   t[8557] := 3_855_850_566;
   t[8558] := 855_950_567;
   t[8559] := 1_856_050_568;
   t[8560] := 2_856_150_569;
   t[8561] := 2_856_250_570;
   t[8562] := 2_856_350_571;
   t[8563] := 1_856_450_572;
   t[8564] := 1_856_550_573;
   t[8565] := 2_856_650_574;
   t[8566] := 2_856_750_575;
   t[8567] := 3_856_850_576;
   t[8568] := 856_950_577;
   t[8569] := 1_857_050_578;
   t[8570] := 1_857_150_579;
   t[8571] := 1_857_250_580;
   t[8572] := 1_857_350_581;
   t[8573] := 2_857_450_582;
   t[8574] := 2_857_550_583;
   t[8575] := 2_857_650_584;
   t[8576] := 3_857_750_585;
   t[8577] := 3_857_850_586;
   t[8578] := 1_857_950_587;
   t[8579] := 1_858_050_588;
   t[8580] := 3_858_150_589;
   t[8581] := 1_858_250_590;
   t[8582] := 3_858_350_591;
   t[8583] := 1_858_450_592;
   t[8584] := 3_858_550_593;
   t[8585] := 858_650_594;
   t[8586] := 858_750_595;
   t[8587] := 1_858_850_596;
   t[8588] := 1_858_950_597;
   t[8589] := 2_859_050_598;
   t[8590] := 1_859_150_599;
   t[8591] := 3_859_250_600;
   t[8592] := 2_859_350_601;
   t[8593] := 859_450_602;
   t[8594] := 859_550_603;
   t[8595] := 1_859_650_604;
   t[8596] := 3_859_750_605;
   t[8597] := 859_850_606;
   t[8598] := 859_950_607;
   t[8599] := 2_860_050_608;
   t[8600] := 3_860_150_609;
   t[8601] := 1_860_250_610;
   t[8602] := 1_860_350_611;
   t[8603] := 2_860_450_612;
   t[8604] := 2_860_550_613;
   t[8605] := 3_860_650_614;
   t[8606] := 3_860_750_615;
   t[8607] := 3_860_850_616;
   t[8608] := 860_950_617;
   t[8609] := 3_861_050_618;
   t[8610] := 861_150_619;
   t[8611] := 861_250_620;
   t[8612] := 2_861_350_621;
   t[8613] := 2_861_450_622;
   t[8614] := 3_861_550_623;
   t[8615] := 2_861_650_624;
   t[8616] := 861_750_625;
   t[8617] := 3_861_850_626;
   t[8618] := 861_950_627;
   t[8619] := 1_862_050_628;
   t[8620] := 1_862_150_629;
   t[8621] := 3_862_250_630;
   t[8622] := 2_862_350_631;
   t[8623] := 3_862_450_632;
   t[8624] := 2_862_550_633;
   t[8625] := 3_862_650_634;
   t[8626] := 3_862_750_635;
   t[8627] := 862_850_636;
   t[8628] := 2_862_950_637;
   t[8629] := 2_863_050_638;
   t[8630] := 863_150_639;
   t[8631] := 3_863_250_640;
   t[8632] := 1_863_350_641;
   t[8633] := 3_863_450_642;
   t[8634] := 3_863_550_643;
   t[8635] := 1_863_650_644;
   t[8636] := 3_863_750_645;
   t[8637] := 1_863_850_646;
   t[8638] := 863_950_647;
   t[8639] := 2_864_050_648;
   t[8640] := 1_864_150_649;
   t[8641] := 2_864_250_650;
   t[8642] := 864_350_651;
   t[8643] := 864_450_652;
   t[8644] := 2_864_550_653;
   t[8645] := 1_864_650_654;
   t[8646] := 3_864_750_655;
   t[8647] := 3_864_850_656;
   t[8648] := 2_864_950_657;
   t[8649] := 865_050_658;
   t[8650] := 1_865_150_659;
   t[8651] := 3_865_250_660;
   t[8652] := 2_865_350_661;
   t[8653] := 865_450_662;
   t[8654] := 3_865_550_663;
   t[8655] := 865_650_664;
   t[8656] := 865_750_665;
   t[8657] := 1_865_850_666;
   t[8658] := 2_865_950_667;
   t[8659] := 3_866_050_668;
   t[8660] := 866_150_669;
   t[8661] := 1_866_250_670;
   t[8662] := 3_866_350_671;
   t[8663] := 2_866_450_672;
   t[8664] := 866_550_673;
   t[8665] := 3_866_650_674;
   t[8666] := 1_866_750_675;
   t[8667] := 1_866_850_676;
   t[8668] := 2_866_950_677;
   t[8669] := 2_867_050_678;
   t[8670] := 3_867_150_679;
   t[8671] := 2_867_250_680;
   t[8672] := 867_350_681;
   t[8673] := 867_450_682;
   t[8674] := 1_867_550_683;
   t[8675] := 867_650_684;
   t[8676] := 2_867_750_685;
   t[8677] := 2_867_850_686;
   t[8678] := 3_867_950_687;
   t[8679] := 3_868_050_688;
   t[8680] := 868_150_689;
   t[8681] := 1_868_250_690;
   t[8682] := 1_868_350_691;
   t[8683] := 2_868_450_692;
   t[8684] := 3_868_550_693;
   t[8685] := 868_650_694;
   t[8686] := 868_750_695;
   t[8687] := 1_868_850_696;
   t[8688] := 2_868_950_697;
   t[8689] := 2_869_050_698;
   t[8690] := 869_150_699;
   t[8691] := 3_869_250_700;
   t[8692] := 1_869_350_701;
   t[8693] := 869_450_702;
   t[8694] := 1_869_550_703;
   t[8695] := 1_869_650_704;
   t[8696] := 2_869_750_705;
   t[8697] := 2_869_850_706;
   t[8698] := 3_869_950_707;
   t[8699] := 3_870_050_708;
   t[8700] := 870_150_709;
   t[8701] := 870_250_710;
   t[8702] := 1_870_350_711;
   t[8703] := 3_870_450_712;
   t[8704] := 3_870_550_713;
   t[8705] := 1_870_650_714;
   t[8706] := 870_750_715;
   t[8707] := 2_870_850_716;
   t[8708] := 2_870_950_717;
   t[8709] := 2_871_050_718;
   t[8710] := 3_871_150_719;
   t[8711] := 3_871_250_720;
   t[8712] := 1_871_350_721;
   t[8713] := 1_871_450_722;
   t[8714] := 2_871_550_723;
   t[8715] := 2_871_650_724;
   t[8716] := 2_871_750_725;
   t[8717] := 1_871_850_726;
   t[8718] := 3_871_950_727;
   t[8719] := 2_872_050_728;
   t[8720] := 872_150_729;
   t[8721] := 872_250_730;
   t[8722] := 1_872_350_731;
   t[8723] := 2_872_450_732;
   t[8724] := 2_872_550_733;
   t[8725] := 872_650_734;
   t[8726] := 3_872_750_735;
   t[8727] := 1_872_850_736;
   t[8728] := 872_950_737;
   t[8729] := 2_873_050_738;
   t[8730] := 2_873_150_739;
   t[8731] := 873_250_740;
   t[8732] := 873_350_741;
   t[8733] := 1_873_450_742;
   t[8734] := 3_873_550_743;
   t[8735] := 873_650_744;
   t[8736] := 2_873_750_745;
   t[8737] := 1_873_850_746;
   t[8738] := 3_873_950_747;
   t[8739] := 2_874_050_748;
   t[8740] := 874_150_749;
   t[8741] := 1_874_250_750;
   t[8742] := 1_874_350_751;
   t[8743] := 3_874_450_752;
   t[8744] := 2_874_550_753;
   t[8745] := 874_650_754;
   t[8746] := 874_750_755;
   t[8747] := 1_874_850_756;
   t[8748] := 2_874_950_757;
   t[8749] := 3_875_050_758;
   t[8750] := 875_150_759;
   t[8751] := 875_250_760;
   t[8752] := 2_875_350_761;
   t[8753] := 2_875_450_762;
   t[8754] := 3_875_550_763;
   t[8755] := 2_875_650_764;
   t[8756] := 875_750_765;
   t[8757] := 1_875_850_766;
   t[8758] := 1_875_950_767;
   t[8759] := 3_876_050_768;
   t[8760] := 876_150_769;
   t[8761] := 1_876_250_770;
   t[8762] := 876_350_771;
   t[8763] := 2_876_450_772;
   t[8764] := 2_876_550_773;
   t[8765] := 876_650_774;
   t[8766] := 3_876_750_775;
   t[8767] := 876_850_776;
   t[8768] := 3_876_950_777;
   t[8769] := 1_877_050_778;
   t[8770] := 1_877_150_779;
   t[8771] := 2_877_250_780;
   t[8772] := 3_877_350_781;
   t[8773] := 877_450_782;
   t[8774] := 2_877_550_783;
   t[8775] := 2_877_650_784;
   t[8776] := 877_750_785;
   t[8777] := 2_877_850_786;
   t[8778] := 877_950_787;
   t[8779] := 3_878_050_788;
   t[8780] := 1_878_150_789;
   t[8781] := 2_878_250_790;
   t[8782] := 2_878_350_791;
   t[8783] := 878_450_792;
   t[8784] := 3_878_550_793;
   t[8785] := 878_650_794;
   t[8786] := 3_878_750_795;
   t[8787] := 1_878_850_796;
   t[8788] := 1_878_950_797;
   t[8789] := 2_879_050_798;
   t[8790] := 3_879_150_799;
   t[8791] := 879_250_800;
   t[8792] := 879_350_801;
   t[8793] := 879_450_802;
   t[8794] := 879_550_803;
   t[8795] := 879_650_804;
   t[8796] := 879_750_805;
   t[8797] := 879_850_806;
   t[8798] := 879_950_807;
   t[8799] := 880_050_808;
   t[8800] := 880_150_809;
   t[8801] := 880_250_810;
   t[8802] := 1_880_350_811;
   t[8803] := 2_880_450_812;
   t[8804] := 3_880_550_813;
   t[8805] := 880_650_814;
   t[8806] := 880_750_815;
   t[8807] := 880_850_816;
   t[8808] := 1_880_950_817;
   t[8809] := 1_881_050_818;
   t[8810] := 3_881_150_819;
   t[8811] := 3_881_250_820;
   t[8812] := 1_881_350_821;
   t[8813] := 2_881_450_822;
   t[8814] := 3_881_550_823;
   t[8815] := 881_650_824;
   t[8816] := 881_750_825;
   t[8817] := 881_850_826;
   t[8818] := 3_881_950_827;
   t[8819] := 3_882_050_828;
   t[8820] := 882_150_829;
   t[8821] := 882_250_830;
   t[8822] := 1_882_350_831;
   t[8823] := 882_450_832;
   t[8824] := 1_882_550_833;
   t[8825] := 1_882_650_834;
   t[8826] := 2_882_750_835;
   t[8827] := 1_882_850_836;
   t[8828] := 3_882_950_837;
   t[8829] := 3_883_050_838;
   t[8830] := 883_150_839;
   t[8831] := 883_250_840;
   t[8832] := 1_883_350_841;
   t[8833] := 2_883_450_842;
   t[8834] := 3_883_550_843;
   t[8835] := 883_650_844;
   t[8836] := 883_750_845;
   t[8837] := 2_883_850_846;
   t[8838] := 2_883_950_847;
   t[8839] := 3_884_050_848;
   t[8840] := 3_884_150_849;
   t[8841] := 1_884_250_850;
   t[8842] := 1_884_350_851;
   t[8843] := 2_884_450_852;
   t[8844] := 1_884_550_853;
   t[8845] := 3_884_650_854;
   t[8846] := 2_884_750_855;
   t[8847] := 884_850_856;
   t[8848] := 884_950_857;
   t[8849] := 2_885_050_858;
   t[8850] := 3_885_150_859;
   t[8851] := 1_885_250_860;
   t[8852] := 1_885_350_861;
   t[8853] := 3_885_450_862;
   t[8854] := 3_885_550_863;
   t[8855] := 885_650_864;
   t[8856] := 1_885_750_865;
   t[8857] := 2_885_850_866;
   t[8858] := 3_885_950_867;
   t[8859] := 886_050_868;
   t[8860] := 886_150_869;
   t[8861] := 886_250_870;
   t[8862] := 886_350_871;
   t[8863] := 1_886_450_872;
   t[8864] := 1_886_550_873;
   t[8865] := 1_886_650_874;
   t[8866] := 1_886_750_875;
   t[8867] := 1_886_850_876;
   t[8868] := 1_886_950_877;
   t[8869] := 887_050_878;
   t[8870] := 887_150_879;
   t[8871] := 2_887_250_880;
   t[8872] := 2_887_350_881;
   t[8873] := 887_450_882;
   t[8874] := 887_550_883;
   t[8875] := 2_887_650_884;
   t[8876] := 1_887_750_885;
   t[8877] := 1_887_850_886;
   t[8878] := 887_950_887;
   t[8879] := 2_888_050_888;
   t[8880] := 2_888_150_889;
   t[8881] := 888_250_890;
   t[8882] := 888_350_891;
   t[8883] := 2_888_450_892;
   t[8884] := 3_888_550_893;
   t[8885] := 3_888_650_894;
   t[8886] := 888_750_895;
   t[8887] := 3_888_850_896;
   t[8888] := 1_888_950_897;
   t[8889] := 1_889_050_898;
   t[8890] := 3_889_150_899;
   t[8891] := 889_250_900;
   t[8892] := 889_350_901;
   t[8893] := 1_889_450_902;
   t[8894] := 2_889_550_903;
   t[8895] := 889_650_904;
   t[8896] := 889_750_905;
   t[8897] := 2_889_850_906;
   t[8898] := 2_889_950_907;
   t[8899] := 890_050_908;
   t[8900] := 3_890_150_909;
   t[8901] := 1_890_250_910;
   t[8902] := 1_890_350_911;
   t[8903] := 2_890_450_912;
   t[8904] := 2_890_550_913;
   t[8905] := 890_650_914;
   t[8906] := 890_750_915;
   t[8907] := 1_890_850_916;
   t[8908] := 1_890_950_917;
   t[8909] := 3_891_050_918;
   t[8910] := 1_891_150_919;
   t[8911] := 3_891_250_920;
   t[8912] := 1_891_350_921;
   t[8913] := 1_891_450_922;
   t[8914] := 3_891_550_923;
   t[8915] := 3_891_650_924;
   t[8916] := 891_750_925;
   t[8917] := 2_891_850_926;
   t[8918] := 1_891_950_927;
   t[8919] := 3_892_050_928;
   t[8920] := 2_892_150_929;
   t[8921] := 3_892_250_930;
   t[8922] := 1_892_350_931;
   t[8923] := 892_450_932;
   t[8924] := 2_892_550_933;
   t[8925] := 2_892_650_934;
   t[8926] := 892_750_935;
   t[8927] := 1_892_850_936;
   t[8928] := 2_892_950_937;
   t[8929] := 893_050_938;
   t[8930] := 893_150_939;
   t[8931] := 2_893_250_940;
   t[8932] := 2_893_350_941;
   t[8933] := 893_450_942;
   t[8934] := 3_893_550_943;
   t[8935] := 1_893_650_944;
   t[8936] := 1_893_750_945;
   t[8937] := 2_893_850_946;
   t[8938] := 2_893_950_947;
   t[8939] := 3_894_050_948;
   t[8940] := 894_150_949;
   t[8941] := 1_894_250_950;
   t[8942] := 2_894_350_951;
   t[8943] := 3_894_450_952;
   t[8944] := 894_550_953;
   t[8945] := 894_650_954;
   t[8946] := 894_750_955;
   t[8947] := 894_850_956;
   t[8948] := 1_894_950_957;
   t[8949] := 1_895_050_958;
   t[8950] := 2_895_150_959;
   t[8951] := 3_895_250_960;
   t[8952] := 895_350_961;
   t[8953] := 895_450_962;
   t[8954] := 3_895_550_963;
   t[8955] := 1_895_650_964;
   t[8956] := 1_895_750_965;
   t[8957] := 3_895_850_966;
   t[8958] := 3_895_950_967;
   t[8959] := 1_896_050_968;
   t[8960] := 1_896_150_969;
   t[8961] := 2_896_250_970;
   t[8962] := 2_896_350_971;
   t[8963] := 3_896_450_972;
   t[8964] := 896_550_973;
   t[8965] := 2_896_650_974;
   t[8966] := 3_896_750_975;
   t[8967] := 1_896_850_976;
   t[8968] := 1_896_950_977;
   t[8969] := 2_897_050_978;
   t[8970] := 3_897_150_979;
   t[8971] := 3_897_250_980;
   t[8972] := 897_350_981;
   t[8973] := 1_897_450_982;
   t[8974] := 2_897_550_983;
   t[8975] := 1_897_650_984;
   t[8976] := 1_897_750_985;
   t[8977] := 1_897_850_986;
   t[8978] := 1_897_950_987;
   t[8979] := 898_050_988;
   t[8980] := 1_898_150_989;
   t[8981] := 1_898_250_990;
   t[8982] := 2_898_350_991;
   t[8983] := 2_898_450_992;
   t[8984] := 898_550_993;
   t[8985] := 898_650_994;
   t[8986] := 2_898_750_995;
   t[8987] := 1_898_850_996;
   t[8988] := 3_898_950_997;
   t[8989] := 2_899_050_998;
   t[8990] := 899_150_999;
   t[8991] := 899_250_001;
   t[8992] := 1_899_350_002;
   t[8993] := 2_899_450_003;
   t[8994] := 3_899_550_004;
   t[8995] := 899_650_005;
   t[8996] := 3_899_750_006;
   t[8997] := 1_899_850_007;
   t[8998] := 899_950_008;
   t[8999] := 1_900_050_009;
   t[9000] := 900_150_010;
   t[9001] := 2_900_250_011;
   t[9002] := 900_350_012;
   t[9003] := 900_450_013;
   t[9004] := 2_900_550_014;
   t[9005] := 1_900_650_015;
   t[9006] := 2_900_750_016;
   t[9007] := 1_900_850_017;
   t[9008] := 3_900_950_018;
   t[9009] := 3_901_050_019;
   t[9010] := 1_901_150_020;
   t[9011] := 1_901_250_021;
   t[9012] := 2_901_350_022;
   t[9013] := 3_901_450_023;
   t[9014] := 2_901_550_024;
   t[9015] := 901_650_025;
   t[9016] := 3_901_750_026;
   t[9017] := 1_901_850_027;
   t[9018] := 1_901_950_028;
   t[9019] := 3_902_050_029;
   t[9020] := 3_902_150_030;
   t[9021] := 902_250_031;
   t[9022] := 3_902_350_032;
   t[9023] := 902_450_033;
   t[9024] := 2_902_550_034;
   t[9025] := 2_902_650_035;
   t[9026] := 902_750_036;
   t[9027] := 902_850_037;
   t[9028] := 2_902_950_038;
   t[9029] := 1_903_050_039;
   t[9030] := 2_903_150_040;
   t[9031] := 1_903_250_041;
   t[9032] := 3_903_350_042;
   t[9033] := 3_903_450_043;
   t[9034] := 903_550_044;
   t[9035] := 1_903_650_045;
   t[9036] := 1_903_750_046;
   t[9037] := 2_903_850_047;
   t[9038] := 2_903_950_048;
   t[9039] := 904_050_049;
   t[9040] := 3_904_150_050;
   t[9041] := 1_904_250_051;
   t[9042] := 904_350_052;
   t[9043] := 2_904_450_053;
   t[9044] := 1_904_550_054;
   t[9045] := 2_904_650_055;
   t[9046] := 1_904_750_056;
   t[9047] := 2_904_850_057;
   t[9048] := 1_904_950_058;
   t[9049] := 3_905_050_059;
   t[9050] := 3_905_150_060;
   t[9051] := 1_905_250_061;
   t[9052] := 1_905_350_062;
   t[9053] := 2_905_450_063;
   t[9054] := 3_905_550_064;
   t[9055] := 905_650_065;
   t[9056] := 905_750_066;
   t[9057] := 1_905_850_067;
   t[9058] := 1_905_950_068;
   t[9059] := 2_906_050_069;
   t[9060] := 2_906_150_070;
   t[9061] := 3_906_250_071;
   t[9062] := 3_906_350_072;
   t[9063] := 3_906_450_073;
   t[9064] := 3_906_550_074;
   t[9065] := 3_906_650_075;
   t[9066] := 3_906_750_076;
   t[9067] := 3_906_850_077;
   t[9068] := 2_906_950_078;
   t[9069] := 2_907_050_079;
   t[9070] := 3_907_150_080;
   t[9071] := 907_250_081;
   t[9072] := 1_907_350_082;
   t[9073] := 2_907_450_083;
   t[9074] := 2_907_550_084;
   t[9075] := 3_907_650_085;
   t[9076] := 3_907_750_086;
   t[9077] := 1_907_850_087;
   t[9078] := 1_907_950_088;
   t[9079] := 3_908_050_089;
   t[9080] := 3_908_150_090;
   t[9081] := 908_250_091;
   t[9082] := 908_350_092;
   t[9083] := 1_908_450_093;
   t[9084] := 2_908_550_094;
   t[9085] := 3_908_650_095;
   t[9086] := 1_908_750_096;
   t[9087] := 2_908_850_097;
   t[9088] := 3_908_950_098;
   t[9089] := 909_050_099;
   t[9090] := 2_909_150_100;
   t[9091] := 909_250_101;
   t[9092] := 2_909_350_102;
   t[9093] := 909_450_103;
   t[9094] := 3_909_550_104;
   t[9095] := 1_909_650_105;
   t[9096] := 1_909_750_106;
   t[9097] := 3_909_850_107;
   t[9098] := 2_909_950_108;
   t[9099] := 3_910_050_109;
   t[9100] := 1_910_150_110;
   t[9101] := 1_910_250_111;
   t[9102] := 3_910_350_112;
   t[9103] := 2_910_450_113;
   t[9104] := 910_550_114;
   t[9105] := 910_650_115;
   t[9106] := 910_750_116;
   t[9107] := 910_850_117;
   t[9108] := 1_910_950_118;
   t[9109] := 3_911_050_119;
   t[9110] := 3_911_150_120;
   t[9111] := 1_911_250_121;
   t[9112] := 1_911_350_122;
   t[9113] := 2_911_450_123;
   t[9114] := 1_911_550_124;
   t[9115] := 2_911_650_125;
   t[9116] := 2_911_750_126;
   t[9117] := 911_850_127;
   t[9118] := 1_911_950_128;
   t[9119] := 2_912_050_129;
   t[9120] := 3_912_150_130;
   t[9121] := 3_912_250_131;
   t[9122] := 1_912_350_132;
   t[9123] := 912_450_133;
   t[9124] := 2_912_550_134;
   t[9125] := 1_912_650_135;
   t[9126] := 3_912_750_136;
   t[9127] := 2_912_850_137;
   t[9128] := 912_950_138;
   t[9129] := 913_050_139;
   t[9130] := 1_913_150_140;
   t[9131] := 3_913_250_141;
   t[9132] := 3_913_350_142;
   t[9133] := 1_913_450_143;
   t[9134] := 913_550_144;
   t[9135] := 2_913_650_145;
   t[9136] := 1_913_750_146;
   t[9137] := 3_913_850_147;
   t[9138] := 913_950_148;
   t[9139] := 1_914_050_149;
   t[9140] := 1_914_150_150;
   t[9141] := 1_914_250_151;
   t[9142] := 2_914_350_152;
   t[9143] := 2_914_450_153;
   t[9144] := 2_914_550_154;
   t[9145] := 1_914_650_155;
   t[9146] := 3_914_750_156;
   t[9147] := 914_850_157;
   t[9148] := 1_914_950_158;
   t[9149] := 1_915_050_159;
   t[9150] := 2_915_150_160;
   t[9151] := 2_915_250_161;
   t[9152] := 3_915_350_162;
   t[9153] := 3_915_450_163;
   t[9154] := 3_915_550_164;
   t[9155] := 3_915_650_165;
   t[9156] := 3_915_750_166;
   t[9157] := 3_915_850_167;
   t[9158] := 3_915_950_168;
   t[9159] := 916_050_169;
   t[9160] := 916_150_170;
   t[9161] := 2_916_250_171;
   t[9162] := 1_916_350_172;
   t[9163] := 3_916_450_173;
   t[9164] := 3_916_550_174;
   t[9165] := 916_650_175;
   t[9166] := 916_750_176;
   t[9167] := 916_850_177;
   t[9168] := 1_916_950_178;
   t[9169] := 1_917_050_179;
   t[9170] := 2_917_150_180;
   t[9171] := 2_917_250_181;
   t[9172] := 3_917_350_182;
   t[9173] := 3_917_450_183;
   t[9174] := 1_917_550_184;
   t[9175] := 3_917_650_185;
   t[9176] := 1_917_750_186;
   t[9177] := 917_850_187;
   t[9178] := 2_917_950_188;
   t[9179] := 1_918_050_189;
   t[9180] := 3_918_150_190;
   t[9181] := 3_918_250_191;
   t[9182] := 918_350_192;
   t[9183] := 918_450_193;
   t[9184] := 1_918_550_194;
   t[9185] := 3_918_650_195;
   t[9186] := 2_918_750_196;
   t[9187] := 918_850_197;
   t[9188] := 918_950_198;
   t[9189] := 2_919_050_199;
   t[9190] := 1_919_150_200;
   t[9191] := 2_919_250_201;
   t[9192] := 3_919_350_202;
   t[9193] := 919_450_203;
   t[9194] := 2_919_550_204;
   t[9195] := 2_919_650_205;
   t[9196] := 919_750_206;
   t[9197] := 3_919_850_207;
   t[9198] := 1_919_950_208;
   t[9199] := 920_050_209;
   t[9200] := 1_920_150_210;
   t[9201] := 2_920_250_211;
   t[9202] := 3_920_350_212;
   t[9203] := 1_920_450_213;
   t[9204] := 1_920_550_214;
   t[9205] := 2_920_650_215;
   t[9206] := 2_920_750_216;
   t[9207] := 920_850_217;
   t[9208] := 3_920_950_218;
   t[9209] := 921_050_219;
   t[9210] := 921_150_220;
   t[9211] := 2_921_250_221;
   t[9212] := 1_921_350_222;
   t[9213] := 2_921_450_223;
   t[9214] := 1_921_550_224;
   t[9215] := 3_921_650_225;
   t[9216] := 3_921_750_226;
   t[9217] := 921_850_227;
   t[9218] := 921_950_228;
   t[9219] := 1_922_050_229;
   t[9220] := 3_922_150_230;
   t[9221] := 3_922_250_231;
   t[9222] := 1_922_350_232;
   t[9223] := 1_922_450_233;
   t[9224] := 3_922_550_234;
   t[9225] := 2_922_650_235;
   t[9226] := 922_750_236;
   t[9227] := 922_850_237;
   t[9228] := 922_950_238;
   t[9229] := 923_050_239;
   t[9230] := 1_923_150_240;
   t[9231] := 2_923_250_241;
   t[9232] := 2_923_350_242;
   t[9233] := 2_923_450_243;
   t[9234] := 2_923_550_244;
   t[9235] := 2_923_650_245;
   t[9236] := 1_923_750_246;
   t[9237] := 2_923_850_247;
   t[9238] := 3_923_950_248;
   t[9239] := 924_050_249;
   t[9240] := 924_150_250;
   t[9241] := 1_924_250_251;
   t[9242] := 2_924_350_252;
   t[9243] := 3_924_450_253;
   t[9244] := 924_550_254;
   t[9245] := 1_924_650_255;
   t[9246] := 2_924_750_256;
   t[9247] := 3_924_850_257;
   t[9248] := 924_950_258;
   t[9249] := 1_925_050_259;
   t[9250] := 2_925_150_260;
   t[9251] := 1_925_250_261;
   t[9252] := 1_925_350_262;
   t[9253] := 1_925_450_263;
   t[9254] := 1_925_550_264;
   t[9255] := 2_925_650_265;
   t[9256] := 2_925_750_266;
   t[9257] := 3_925_850_267;
   t[9258] := 3_925_950_268;
   t[9259] := 3_926_050_269;
   t[9260] := 3_926_150_270;
   t[9261] := 1_926_250_271;
   t[9262] := 2_926_350_272;
   t[9263] := 3_926_450_273;
   t[9264] := 3_926_550_274;
   t[9265] := 926_650_275;
   t[9266] := 926_750_276;
   t[9267] := 1_926_850_277;
   t[9268] := 1_926_950_278;
   t[9269] := 2_927_050_279;
   t[9270] := 2_927_150_280;
   t[9271] := 3_927_250_281;
   t[9272] := 927_350_282;
   t[9273] := 927_450_283;
   t[9274] := 927_550_284;
   t[9275] := 1_927_650_285;
   t[9276] := 2_927_750_286;
   t[9277] := 2_927_850_287;
   t[9278] := 927_950_288;
   t[9279] := 928_050_289;
   t[9280] := 2_928_150_290;
   t[9281] := 2_928_250_291;
   t[9282] := 3_928_350_292;
   t[9283] := 928_450_293;
   t[9284] := 1_928_550_294;
   t[9285] := 1_928_650_295;
   t[9286] := 2_928_750_296;
   t[9287] := 2_928_850_297;
   t[9288] := 3_928_950_298;
   t[9289] := 3_929_050_299;
   t[9290] := 929_150_300;
   t[9291] := 929_250_301;
   t[9292] := 1_929_350_302;
   t[9293] := 1_929_450_303;
   t[9294] := 2_929_550_304;
   t[9295] := 3_929_650_305;
   t[9296] := 3_929_750_306;
   t[9297] := 929_850_307;
   t[9298] := 929_950_308;
   t[9299] := 2_930_050_309;
   t[9300] := 1_930_150_310;
   t[9301] := 3_930_250_311;
   t[9302] := 2_930_350_312;
   t[9303] := 930_450_313;
   t[9304] := 1_930_550_314;
   t[9305] := 1_930_650_315;
   t[9306] := 3_930_750_316;
   t[9307] := 2_930_850_317;
   t[9308] := 930_950_318;
   t[9309] := 1_931_050_319;
   t[9310] := 2_931_150_320;
   t[9311] := 3_931_250_321;
   t[9312] := 3_931_350_322;
   t[9313] := 931_450_323;
   t[9314] := 1_931_550_324;
   t[9315] := 2_931_650_325;
   t[9316] := 2_931_750_326;
   t[9317] := 931_850_327;
   t[9318] := 3_931_950_328;
   t[9319] := 1_932_050_329;
   t[9320] := 932_150_330;
   t[9321] := 2_932_250_331;
   t[9322] := 2_932_350_332;
   t[9323] := 3_932_450_333;
   t[9324] := 932_550_334;
   t[9325] := 1_932_650_335;
   t[9326] := 2_932_750_336;
   t[9327] := 1_932_850_337;
   t[9328] := 2_932_950_338;
   t[9329] := 2_933_050_339;
   t[9330] := 933_150_340;
   t[9331] := 933_250_341;
   t[9332] := 2_933_350_342;
   t[9333] := 3_933_450_343;
   t[9334] := 1_933_550_344;
   t[9335] := 933_650_345;
   t[9336] := 2_933_750_346;
   t[9337] := 933_850_347;
   t[9338] := 2_933_950_348;
   t[9339] := 934_050_349;
   t[9340] := 1_934_150_350;
   t[9341] := 2_934_250_351;
   t[9342] := 2_934_350_352;
   t[9343] := 2_934_450_353;
   t[9344] := 2_934_550_354;
   t[9345] := 2_934_650_355;
   t[9346] := 3_934_750_356;
   t[9347] := 3_934_850_357;
   t[9348] := 934_950_358;
   t[9349] := 1_935_050_359;
   t[9350] := 1_935_150_360;
   t[9351] := 2_935_250_361;
   t[9352] := 3_935_350_362;
   t[9353] := 3_935_450_363;
   t[9354] := 935_550_364;
   t[9355] := 1_935_650_365;
   t[9356] := 2_935_750_366;
   t[9357] := 3_935_850_367;
   t[9358] := 3_935_950_368;
   t[9359] := 3_936_050_369;
   t[9360] := 3_936_150_370;
   t[9361] := 3_936_250_371;
   t[9362] := 936_350_372;
   t[9363] := 1_936_450_373;
   t[9364] := 1_936_550_374;
   t[9365] := 3_936_650_375;
   t[9366] := 3_936_750_376;
   t[9367] := 1_936_850_377;
   t[9368] := 936_950_378;
   t[9369] := 2_937_050_379;
   t[9370] := 2_937_150_380;
   t[9371] := 937_250_381;
   t[9372] := 937_350_382;
   t[9373] := 1_937_450_383;
   t[9374] := 1_937_550_384;
   t[9375] := 2_937_650_385;
   t[9376] := 3_937_750_386;
   t[9377] := 937_850_387;
   t[9378] := 1_937_950_388;
   t[9379] := 1_938_050_389;
   t[9380] := 3_938_150_390;
   t[9381] := 1_938_250_391;
   t[9382] := 3_938_350_392;
   t[9383] := 3_938_450_393;
   t[9384] := 1_938_550_394;
   t[9385] := 3_938_650_395;
   t[9386] := 3_938_750_396;
   t[9387] := 1_938_850_397;
   t[9388] := 3_938_950_398;
   t[9389] := 1_939_050_399;
   t[9390] := 939_150_400;
   t[9391] := 2_939_250_401;
   t[9392] := 2_939_350_402;
   t[9393] := 939_450_403;
   t[9394] := 2_939_550_404;
   t[9395] := 1_939_650_405;
   t[9396] := 2_939_750_406;
   t[9397] := 2_939_850_407;
   t[9398] := 3_939_950_408;
   t[9399] := 3_940_050_409;
   t[9400] := 1_940_150_410;
   t[9401] := 940_250_411;
   t[9402] := 2_940_350_412;
   t[9403] := 2_940_450_413;
   t[9404] := 2_940_550_414;
   t[9405] := 2_940_650_415;
   t[9406] := 3_940_750_416;
   t[9407] := 940_850_417;
   t[9408] := 1_940_950_418;
   t[9409] := 2_941_050_419;
   t[9410] := 3_941_150_420;
   t[9411] := 941_250_421;
   t[9412] := 3_941_350_422;
   t[9413] := 1_941_450_423;
   t[9414] := 941_550_424;
   t[9415] := 2_941_650_425;
   t[9416] := 1_941_750_426;
   t[9417] := 3_941_850_427;
   t[9418] := 941_950_428;
   t[9419] := 942_050_429;
   t[9420] := 2_942_150_430;
   t[9421] := 1_942_250_431;
   t[9422] := 3_942_350_432;
   t[9423] := 2_942_450_433;
   t[9424] := 942_550_434;
   t[9425] := 942_650_435;
   t[9426] := 1_942_750_436;
   t[9427] := 1_942_850_437;
   t[9428] := 1_942_950_438;
   t[9429] := 2_943_050_439;
   t[9430] := 1_943_150_440;
   t[9431] := 3_943_250_441;
   t[9432] := 3_943_350_442;
   t[9433] := 1_943_450_443;
   t[9434] := 2_943_550_444;
   t[9435] := 2_943_650_445;
   t[9436] := 943_750_446;
   t[9437] := 3_943_850_447;
   t[9438] := 1_943_950_448;
   t[9439] := 944_050_449;
   t[9440] := 2_944_150_450;
   t[9441] := 2_944_250_451;
   t[9442] := 3_944_350_452;
   t[9443] := 944_450_453;
   t[9444] := 1_944_550_454;
   t[9445] := 3_944_650_455;
   t[9446] := 2_944_750_456;
   t[9447] := 944_850_457;
   t[9448] := 1_944_950_458;
   t[9449] := 2_945_050_459;
   t[9450] := 3_945_150_460;
   t[9451] := 3_945_250_461;
   t[9452] := 1_945_350_462;
   t[9453] := 945_450_463;
   t[9454] := 2_945_550_464;
   t[9455] := 1_945_650_465;
   t[9456] := 3_945_750_466;
   t[9457] := 3_945_850_467;
   t[9458] := 3_945_950_468;
   t[9459] := 1_946_050_469;
   t[9460] := 946_150_470;
   t[9461] := 2_946_250_471;
   t[9462] := 1_946_350_472;
   t[9463] := 2_946_450_473;
   t[9464] := 2_946_550_474;
   t[9465] := 2_946_650_475;
   t[9466] := 2_946_750_476;
   t[9467] := 3_946_850_477;
   t[9468] := 3_946_950_478;
   t[9469] := 947_050_479;
   t[9470] := 1_947_150_480;
   t[9471] := 2_947_250_481;
   t[9472] := 2_947_350_482;
   t[9473] := 2_947_450_483;
   t[9474] := 2_947_550_484;
   t[9475] := 2_947_650_485;
   t[9476] := 2_947_750_486;
   t[9477] := 3_947_850_487;
   t[9478] := 3_947_950_488;
   t[9479] := 948_050_489;
   t[9480] := 948_150_490;
   t[9481] := 948_250_491;
   t[9482] := 1_948_350_492;
   t[9483] := 1_948_450_493;
   t[9484] := 2_948_550_494;
   t[9485] := 3_948_650_495;
   t[9486] := 3_948_750_496;
   t[9487] := 1_948_850_497;
   t[9488] := 948_950_498;
   t[9489] := 1_949_050_499;
   t[9490] := 2_949_150_500;
   t[9491] := 2_949_250_501;
   t[9492] := 3_949_350_502;
   t[9493] := 1_949_450_503;
   t[9494] := 1_949_550_504;
   t[9495] := 3_949_650_505;
   t[9496] := 1_949_750_506;
   t[9497] := 2_949_850_507;
   t[9498] := 1_949_950_508;
   t[9499] := 3_950_050_509;
   t[9500] := 1_950_150_510;
   t[9501] := 1_950_250_511;
   t[9502] := 3_950_350_512;
   t[9503] := 2_950_450_513;
   t[9504] := 950_550_514;
   t[9505] := 950_650_515;
   t[9506] := 1_950_750_516;
   t[9507] := 1_950_850_517;
   t[9508] := 3_950_950_518;
   t[9509] := 3_951_050_519;
   t[9510] := 951_150_520;
   t[9511] := 3_951_250_521;
   t[9512] := 951_350_522;
   t[9513] := 1_951_450_523;
   t[9514] := 2_951_550_524;
   t[9515] := 3_951_650_525;
   t[9516] := 3_951_750_526;
   t[9517] := 1_951_850_527;
   t[9518] := 951_950_528;
   t[9519] := 2_952_050_529;
   t[9520] := 1_952_150_530;
   t[9521] := 3_952_250_531;
   t[9522] := 3_952_350_532;
   t[9523] := 952_450_533;
   t[9524] := 1_952_550_534;
   t[9525] := 2_952_650_535;
   t[9526] := 3_952_750_536;
   t[9527] := 2_952_850_537;
   t[9528] := 952_950_538;
   t[9529] := 3_953_050_539;
   t[9530] := 1_953_150_540;
   t[9531] := 1_953_250_541;
   t[9532] := 2_953_350_542;
   t[9533] := 953_450_543;
   t[9534] := 3_953_550_544;
   t[9535] := 1_953_650_545;
   t[9536] := 953_750_546;
   t[9537] := 2_953_850_547;
   t[9538] := 2_953_950_548;
   t[9539] := 954_050_549;
   t[9540] := 954_150_550;
   t[9541] := 954_250_551;
   t[9542] := 954_350_552;
   t[9543] := 954_450_553;
   t[9544] := 1_954_550_554;
   t[9545] := 3_954_650_555;
   t[9546] := 954_750_556;
   t[9547] := 1_954_850_557;
   t[9548] := 2_954_950_558;
   t[9549] := 1_955_050_559;
   t[9550] := 3_955_150_560;
   t[9551] := 1_955_250_561;
   t[9552] := 3_955_350_562;
   t[9553] := 2_955_450_563;
   t[9554] := 955_550_564;
   t[9555] := 955_650_565;
   t[9556] := 2_955_750_566;
   t[9557] := 1_955_850_567;
   t[9558] := 1_955_950_568;
   t[9559] := 3_956_050_569;
   t[9560] := 2_956_150_570;
   t[9561] := 956_250_571;
   t[9562] := 1_956_350_572;
   t[9563] := 1_956_450_573;
   t[9564] := 3_956_550_574;
   t[9565] := 956_650_575;
   t[9566] := 2_956_750_576;
   t[9567] := 956_850_577;
   t[9568] := 2_956_950_578;
   t[9569] := 957_050_579;
   t[9570] := 2_957_150_580;
   t[9571] := 957_250_581;
   t[9572] := 2_957_350_582;
   t[9573] := 2_957_450_583;
   t[9574] := 2_957_550_584;
   t[9575] := 957_650_585;
   t[9576] := 3_957_750_586;
   t[9577] := 1_957_850_587;
   t[9578] := 1_957_950_588;
   t[9579] := 3_958_050_589;
   t[9580] := 958_150_590;
   t[9581] := 3_958_250_591;
   t[9582] := 1_958_350_592;
   t[9583] := 3_958_450_593;
   t[9584] := 1_958_550_594;
   t[9585] := 3_958_650_595;
   t[9586] := 3_958_750_596;
   t[9587] := 1_958_850_597;
   t[9588] := 958_950_598;
   t[9589] := 2_959_050_599;
   t[9590] := 2_959_150_600;
   t[9591] := 2_959_250_601;
   t[9592] := 959_350_602;
   t[9593] := 959_450_603;
   t[9594] := 2_959_550_604;
   t[9595] := 1_959_650_605;
   t[9596] := 3_959_750_606;
   t[9597] := 959_850_607;
   t[9598] := 959_950_608;
   t[9599] := 2_960_050_609;
   t[9600] := 2_960_150_610;
   t[9601] := 3_960_250_611;
   t[9602] := 960_350_612;
   t[9603] := 1_960_450_613;
   t[9604] := 960_550_614;
   t[9605] := 2_960_650_615;
   t[9606] := 960_750_616;
   t[9607] := 3_960_850_617;
   t[9608] := 960_950_618;
   t[9609] := 961_050_619;
   t[9610] := 2_961_150_620;
   t[9611] := 3_961_250_621;
   t[9612] := 2_961_350_622;
   t[9613] := 961_450_623;
   t[9614] := 961_550_624;
   t[9615] := 1_961_650_625;
   t[9616] := 2_961_750_626;
   t[9617] := 2_961_850_627;
   t[9618] := 961_950_628;
   t[9619] := 3_962_050_629;
   t[9620] := 1_962_150_630;
   t[9621] := 962_250_631;
   t[9622] := 2_962_350_632;
   t[9623] := 2_962_450_633;
   t[9624] := 3_962_550_634;
   t[9625] := 1_962_650_635;
   t[9626] := 962_750_636;
   t[9627] := 2_962_850_637;
   t[9628] := 1_962_950_638;
   t[9629] := 3_963_050_639;
   t[9630] := 963_150_640;
   t[9631] := 1_963_250_641;
   t[9632] := 2_963_350_642;
   t[9633] := 2_963_450_643;
   t[9634] := 1_963_550_644;
   t[9635] := 1_963_650_645;
   t[9636] := 3_963_750_646;
   t[9637] := 3_963_850_647;
   t[9638] := 1_963_950_648;
   t[9639] := 1_964_050_649;
   t[9640] := 3_964_150_650;
   t[9641] := 3_964_250_651;
   t[9642] := 964_350_652;
   t[9643] := 3_964_450_653;
   t[9644] := 1_964_550_654;
   t[9645] := 1_964_650_655;
   t[9646] := 3_964_750_656;
   t[9647] := 3_964_850_657;
   t[9648] := 1_964_950_658;
   t[9649] := 1_965_050_659;
   t[9650] := 2_965_150_660;
   t[9651] := 965_250_661;
   t[9652] := 1_965_350_662;
   t[9653] := 1_965_450_663;
   t[9654] := 3_965_550_664;
   t[9655] := 3_965_650_665;
   t[9656] := 965_750_666;
   t[9657] := 2_965_850_667;
   t[9658] := 965_950_668;
   t[9659] := 966_050_669;
   t[9660] := 1_966_150_670;
   t[9661] := 2_966_250_671;
   t[9662] := 2_966_350_672;
   t[9663] := 3_966_450_673;
   t[9664] := 2_966_550_674;
   t[9665] := 3_966_650_675;
   t[9666] := 3_966_750_676;
   t[9667] := 1_966_850_677;
   t[9668] := 966_950_678;
   t[9669] := 2_967_050_679;
   t[9670] := 2_967_150_680;
   t[9671] := 3_967_250_681;
   t[9672] := 3_967_350_682;
   t[9673] := 3_967_450_683;
   t[9674] := 3_967_550_684;
   t[9675] := 3_967_650_685;
   t[9676] := 967_750_686;
   t[9677] := 967_850_687;
   t[9678] := 2_967_950_688;
   t[9679] := 2_968_050_689;
   t[9680] := 3_968_150_690;
   t[9681] := 3_968_250_691;
   t[9682] := 1_968_350_692;
   t[9683] := 1_968_450_693;
   t[9684] := 3_968_550_694;
   t[9685] := 2_968_650_695;
   t[9686] := 3_968_750_696;
   t[9687] := 3_968_850_697;
   t[9688] := 968_950_698;
   t[9689] := 1_969_050_699;
   t[9690] := 2_969_150_700;
   t[9691] := 2_969_250_701;
   t[9692] := 2_969_350_702;
   t[9693] := 3_969_450_703;
   t[9694] := 2_969_550_704;
   t[9695] := 3_969_650_705;
   t[9696] := 2_969_750_706;
   t[9697] := 969_850_707;
   t[9698] := 1_969_950_708;
   t[9699] := 2_970_050_709;
   t[9700] := 970_150_710;
   t[9701] := 970_250_711;
   t[9702] := 2_970_350_712;
   t[9703] := 970_450_713;
   t[9704] := 2_970_550_714;
   t[9705] := 2_970_650_715;
   t[9706] := 970_750_716;
   t[9707] := 1_970_850_717;
   t[9708] := 1_970_950_718;
   t[9709] := 3_971_050_719;
   t[9710] := 1_971_150_720;
   t[9711] := 3_971_250_721;
   t[9712] := 2_971_350_722;
   t[9713] := 971_450_723;
   t[9714] := 971_550_724;
   t[9715] := 2_971_650_725;
   t[9716] := 3_971_750_726;
   t[9717] := 971_850_727;
   t[9718] := 971_950_728;
   t[9719] := 3_972_050_729;
   t[9720] := 1_972_150_730;
   t[9721] := 972_250_731;
   t[9722] := 2_972_350_732;
   t[9723] := 1_972_450_733;
   t[9724] := 3_972_550_734;
   t[9725] := 2_972_650_735;
   t[9726] := 3_972_750_736;
   t[9727] := 2_972_850_737;
   t[9728] := 972_950_738;
   t[9729] := 973_050_739;
   t[9730] := 2_973_150_740;
   t[9731] := 2_973_250_741;
   t[9732] := 973_350_742;
   t[9733] := 3_973_450_743;
   t[9734] := 973_550_744;
   t[9735] := 1_973_650_745;
   t[9736] := 1_973_750_746;
   t[9737] := 2_973_850_747;
   t[9738] := 2_973_950_748;
   t[9739] := 3_974_050_749;
   t[9740] := 974_150_750;
   t[9741] := 974_250_751;
   t[9742] := 1_974_350_752;
   t[9743] := 3_974_450_753;
   t[9744] := 3_974_550_754;
   t[9745] := 1_974_650_755;
   t[9746] := 2_974_750_756;
   t[9747] := 3_974_850_757;
   t[9748] := 974_950_758;
   t[9749] := 1_975_050_759;
   t[9750] := 2_975_150_760;
   t[9751] := 2_975_250_761;
   t[9752] := 2_975_350_762;
   t[9753] := 2_975_450_763;
   t[9754] := 2_975_550_764;
   t[9755] := 2_975_650_765;
   t[9756] := 1_975_750_766;
   t[9757] := 1_975_850_767;
   t[9758] := 2_975_950_768;
   t[9759] := 2_976_050_769;
   t[9760] := 976_150_770;
   t[9761] := 3_976_250_771;
   t[9762] := 976_350_772;
   t[9763] := 976_450_773;
   t[9764] := 1_976_550_774;
   t[9765] := 1_976_650_775;
   t[9766] := 3_976_750_776;
   t[9767] := 3_976_850_777;
   t[9768] := 976_950_778;
   t[9769] := 1_977_050_779;
   t[9770] := 2_977_150_780;
   t[9771] := 2_977_250_781;
   t[9772] := 2_977_350_782;
   t[9773] := 2_977_450_783;
   t[9774] := 3_977_550_784;
   t[9775] := 3_977_650_785;
   t[9776] := 3_977_750_786;
   t[9777] := 977_850_787;
   t[9778] := 1_977_950_788;
   t[9779] := 1_978_050_789;
   t[9780] := 3_978_150_790;
   t[9781] := 978_250_791;
   t[9782] := 2_978_350_792;
   t[9783] := 3_978_450_793;
   t[9784] := 3_978_550_794;
   t[9785] := 978_650_795;
   t[9786] := 1_978_750_796;
   t[9787] := 3_978_850_797;
   t[9788] := 3_978_950_798;
   t[9789] := 1_979_050_799;
   t[9790] := 1_979_150_800;
   t[9791] := 3_979_250_801;
   t[9792] := 2_979_350_802;
   t[9793] := 979_450_803;
   t[9794] := 979_550_804;
   t[9795] := 1_979_650_805;
   t[9796] := 1_979_750_806;
   t[9797] := 3_979_850_807;
   t[9798] := 2_979_950_808;
   t[9799] := 980_050_809;
   t[9800] := 1_980_150_810;
   t[9801] := 2_980_250_811;
   t[9802] := 3_980_350_812;
   t[9803] := 2_980_450_813;
   t[9804] := 3_980_550_814;
   t[9805] := 2_980_650_815;
   t[9806] := 980_750_816;
   t[9807] := 1_980_850_817;
   t[9808] := 2_980_950_818;
   t[9809] := 981_050_819;
   t[9810] := 1_981_150_820;
   t[9811] := 1_981_250_821;
   t[9812] := 3_981_350_822;
   t[9813] := 2_981_450_823;
   t[9814] := 981_550_824;
   t[9815] := 981_650_825;
   t[9816] := 2_981_750_826;
   t[9817] := 3_981_850_827;
   t[9818] := 3_981_950_828;
   t[9819] := 1_982_050_829;
   t[9820] := 1_982_150_830;
   t[9821] := 2_982_250_831;
   t[9822] := 3_982_350_832;
   t[9823] := 982_450_833;
   t[9824] := 2_982_550_834;
   t[9825] := 2_982_650_835;
   t[9826] := 3_982_750_836;
   t[9827] := 2_982_850_837;
   t[9828] := 982_950_838;
   t[9829] := 983_050_839;
   t[9830] := 2_983_150_840;
   t[9831] := 3_983_250_841;
   t[9832] := 983_350_842;
   t[9833] := 1_983_450_843;
   t[9834] := 1_983_550_844;
   t[9835] := 3_983_650_845;
   t[9836] := 1_983_750_846;
   t[9837] := 983_850_847;
   t[9838] := 1_983_950_848;
   t[9839] := 2_984_050_849;
   t[9840] := 3_984_150_850;
   t[9841] := 984_250_851;
   t[9842] := 984_350_852;
   t[9843] := 2_984_450_853;
   t[9844] := 2_984_550_854;
   t[9845] := 984_650_855;
   t[9846] := 3_984_750_856;
   t[9847] := 1_984_850_857;
   t[9848] := 984_950_858;
   t[9849] := 2_985_050_859;
   t[9850] := 2_985_150_860;
   t[9851] := 3_985_250_861;
   t[9852] := 3_985_350_862;
   t[9853] := 985_450_863;
   t[9854] := 985_550_864;
   t[9855] := 1_985_650_865;
   t[9856] := 1_985_750_866;
   t[9857] := 3_985_850_867;
   t[9858] := 985_950_868;
   t[9859] := 1_986_050_869;
   t[9860] := 1_986_150_870;
   t[9861] := 1_986_250_871;
   t[9862] := 3_986_350_872;
   t[9863] := 2_986_450_873;
   t[9864] := 3_986_550_874;
   t[9865] := 986_650_875;
   t[9866] := 2_986_750_876;
   t[9867] := 3_986_850_877;
   t[9868] := 1_986_950_878;
   t[9869] := 2_987_050_879;
   t[9870] := 3_987_150_880;
   t[9871] := 3_987_250_881;
   t[9872] := 3_987_350_882;
   t[9873] := 3_987_450_883;
   t[9874] := 987_550_884;
   t[9875] := 987_650_885;
   t[9876] := 2_987_750_886;
   t[9877] := 2_987_850_887;
   t[9878] := 987_950_888;
   t[9879] := 3_988_050_889;
   t[9880] := 2_988_150_890;
   t[9881] := 3_988_250_891;
   t[9882] := 1_988_350_892;
   t[9883] := 2_988_450_893;
   t[9884] := 2_988_550_894;
   t[9885] := 988_650_895;
   t[9886] := 1_988_750_896;
   t[9887] := 1_988_850_897;
   t[9888] := 3_988_950_898;
   t[9889] := 1_989_050_899;
   t[9890] := 3_989_150_900;
   t[9891] := 3_989_250_901;
   t[9892] := 1_989_350_902;
   t[9893] := 1_989_450_903;
   t[9894] := 2_989_550_904;
   t[9895] := 2_989_650_905;
   t[9896] := 3_989_750_906;
   t[9897] := 3_989_850_907;
   t[9898] := 2_989_950_908;
   t[9899] := 990_050_909;
   t[9900] := 2_990_150_910;
   t[9901] := 990_250_911;
   t[9902] := 1_990_350_912;
   t[9903] := 1_990_450_913;
   t[9904] := 3_990_550_914;
   t[9905] := 990_650_915;
   t[9906] := 990_750_916;
   t[9907] := 2_990_850_917;
   t[9908] := 1_990_950_918;
   t[9909] := 2_991_050_919;
   t[9910] := 1_991_150_920;
   t[9911] := 3_991_250_921;
   t[9912] := 3_991_350_922;
   t[9913] := 991_450_923;
   t[9914] := 991_550_924;
   t[9915] := 991_650_925;
   t[9916] := 2_991_750_926;
   t[9917] := 991_850_927;
   t[9918] := 2_991_950_928;
   t[9919] := 3_992_050_929;
   t[9920] := 992_150_930;
   t[9921] := 2_992_250_931;
   t[9922] := 3_992_350_932;
   t[9923] := 1_992_450_933;
   t[9924] := 992_550_934;
   t[9925] := 2_992_650_935;
   t[9926] := 1_992_750_936;
   t[9927] := 3_992_850_937;
   t[9928] := 2_992_950_938;
   t[9929] := 993_050_939;
   t[9930] := 993_150_940;
   t[9931] := 1_993_250_941;
   t[9932] := 2_993_350_942;
   t[9933] := 3_993_450_943;
   t[9934] := 1_993_550_944;
   t[9935] := 1_993_650_945;
   t[9936] := 3_993_750_946;
   t[9937] := 2_993_850_947;
   t[9938] := 993_950_948;
   t[9939] := 3_994_050_949;
   t[9940] := 994_150_950;
   t[9941] := 994_250_951;
   t[9942] := 1_994_350_952;
   t[9943] := 994_450_953;
   t[9944] := 2_994_550_954;
   t[9945] := 994_650_955;
   t[9946] := 2_994_750_956;
   t[9947] := 994_850_957;
   t[9948] := 2_994_950_958;
   t[9949] := 3_995_050_959;
   t[9950] := 995_150_960;
   t[9951] := 1_995_250_961;
   t[9952] := 3_995_350_962;
   t[9953] := 995_450_963;
   t[9954] := 2_995_550_964;
   t[9955] := 3_995_650_965;
   t[9956] := 1_995_750_966;
   t[9957] := 3_995_850_967;
   t[9958] := 1_995_950_968;
   t[9959] := 3_996_050_969;
   t[9960] := 1_996_150_970;
   t[9961] := 3_996_250_971;
   t[9962] := 1_996_350_972;
   t[9963] := 3_996_450_973;
   t[9964] := 2_996_550_974;
   t[9965] := 996_650_975;
   t[9966] := 2_996_750_976;
   t[9967] := 996_850_977;
   t[9968] := 2_996_950_978;
   t[9969] := 997_050_979;
   t[9970] := 2_997_150_980;
   t[9971] := 3_997_250_981;
   t[9972] := 997_350_982;
   t[9973] := 1_997_450_983;
   t[9974] := 2_997_550_984;
   t[9975] := 3_997_650_985;
   t[9976] := 997_750_986;
   t[9977] := 1_997_850_987;
   t[9978] := 2_997_950_988;
   t[9979] := 3_998_050_989;
   t[9980] := 998_150_990;
   t[9981] := 1_998_250_991;
   t[9982] := 2_998_350_992;
   t[9983] := 2_998_450_993;
   t[9984] := 998_550_994;
   t[9985] := 1_998_650_995;
   t[9986] := 2_998_750_996;
   t[9987] := 998_850_997;
   t[9988] := 1_998_950_998;
   t[9989] := 2_999_050_999;
   t[9990] := 3_999_150_001;
   t[9991] := 999_250_002;
   t[9992] := 1_999_350_003;
   t[9993] := 1_999_450_004;
   t[9994] := 3_999_550_005;
   t[9995] := 1_999_650_006;
   t[9996] := 2_999_750_007;
   t[9997] := 999_850_008;
   t[9998] := 0;
   t[9999] := 0;
   t[10000] := 0;
END_DATA_BLOCK

// folder: (top level)

FUNCTION_BLOCK "FB1_DRIVE"   // FB1, LAD
{ S7_Optimized_Access := 'TRUE' }
VERSION : 0.1
   VAR_INPUT
      iStart : Bool;
      iStop : Bool;
      iProtectie : Bool;
      iContactor : Bool;
      iBrake : Bool;
      iRun : Bool;
      iFault : Bool;
      iResetFault : Bool;
      iAck_Fault : Bool;
   END_VAR
   VAR_OUTPUT
      oContactor : Bool;
      oON : Bool;
      oBrake : Bool;
      oFault : Bool;
      oAlarmProtectie : Bool;
      oAlarmContactor : Bool;
      oAlarmBrake : Bool;
      oBlocked : Bool;
      oFaultBrake : Bool;
      oFaultContactor : Bool;
      oAckFault : Bool;
   END_VAR
   VAR
      Release_Brake : Bool;
      Cuplare : Bool;
   END_VAR
BEGIN

REGION Network 1
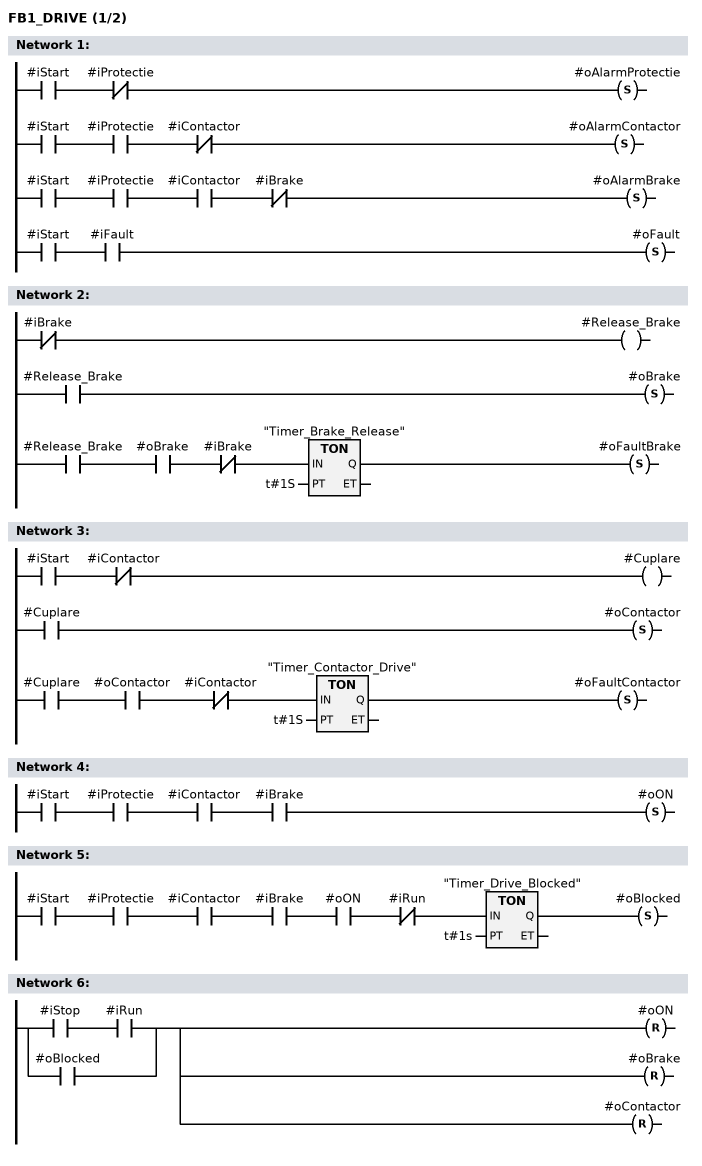
   RUNG wire#powerrail
      Contact( #iStart )
      I_Contact( #iProtectie )
      S_Coil( #oAlarmProtectie )
   END_RUNG
   RUNG wire#powerrail
      Contact( #iStart )
      Contact( #iProtectie )
      I_Contact( #iContactor )
      S_Coil( #oAlarmContactor )
   END_RUNG
   RUNG wire#powerrail
      Contact( #iStart )
      Contact( #iProtectie )
      Contact( #iContactor )
      I_Contact( #iBrake )
      S_Coil( #oAlarmBrake )
   END_RUNG
   RUNG wire#powerrail
      Contact( #iStart )
      Contact( #iFault )
      S_Coil( #oFault )
   END_RUNG
   // the same network as SCL:
   IF #iStart AND NOT #iProtectie THEN #oAlarmProtectie := TRUE; END_IF;
   IF #iStart AND #iProtectie AND NOT #iContactor THEN #oAlarmContactor := TRUE; END_IF;
   IF #iStart AND #iProtectie AND #iContactor AND NOT #iBrake THEN #oAlarmBrake := TRUE; END_IF;
   IF #iStart AND #iFault THEN #oFault := TRUE; END_IF;
END_REGION

REGION Network 2
   #Release_Brake := NOT #iBrake;
   IF #Release_Brake THEN #oBrake := TRUE; END_IF;
   "Timer_Brake_Release".TON(IN := #Release_Brake AND #oBrake AND NOT #iBrake, PT := t#1S);
   IF "Timer_Brake_Release".Q THEN #oFaultBrake := TRUE; END_IF;
END_REGION

REGION Network 3
   #Cuplare := #iStart AND NOT #iContactor;
   IF #Cuplare THEN #oContactor := TRUE; END_IF;
   "Timer_Contactor_Drive".TON(IN := #Cuplare AND #oContactor AND NOT #iContactor, PT := t#1S);
   IF "Timer_Contactor_Drive".Q THEN #oFaultContactor := TRUE; END_IF;
END_REGION

REGION Network 4
   RUNG wire#powerrail
      Contact( #iStart )
      Contact( #iProtectie )
      Contact( #iContactor )
      Contact( #iBrake )
      S_Coil( #oON )
   END_RUNG
   // the same network as SCL:
   IF #iStart AND #iProtectie AND #iContactor AND #iBrake THEN #oON := TRUE; END_IF;
END_REGION

REGION Network 5
   "Timer_Drive_Blocked".TON(IN := #iStart AND #iProtectie AND #iContactor AND #iBrake AND #oON AND NOT #iRun,
                           PT := t#1s);
   IF "Timer_Drive_Blocked".Q THEN #oBlocked := TRUE; END_IF;
END_REGION
